FUNCTION "FC116_Inerting" : Void   // FC116, STL
{ S7_Optimized_Access := 'FALSE' }
AUTHOR : JaegerA
FAMILY : RS_KK
NAME : Inerting
VERSION : 1.1
   VAR_INPUT
      IN_Enable : Bool;
      IN_With_Inerting : Bool;   // Inerting selected in TP
      IN_OP_Mode_Manual : Bool;
      IN_OP_Mode_Wetshot : Bool;
      IN_OP_Mode_Test : Bool;
      IN_Start : Bool;
      IN_Stop : Bool;
      IN_T_Flushing : Bool;
      IN_T_Purge_Air : Bool;
      IN_Enable_pressurize_time : Bool;
      IN_AutoPurge_Air : Bool;
      IN_Quitt_Fault : Bool;
      IN_Cycle_runs : Bool;
      IN_MC_Activ : Bool;
      IN_PressurizeTimeRuns : Bool;
      IN_Shotend : Bool;
      IN_S_P_N2 : Bool;
      IN_S_P_FlushingAgent : Bool;
      IN_MH_selected : Bool;
      IN_Inert_MH : Bool;
      IN_Inert_Lance : Bool;
      IN_IntervalCleaning : Bool;
      IN_Ctrl_Fault_On : Bool;
      IN_Flowrate_N2_Actual : Real;
      IN_Shotwight : Real;
      IN_Foam_Density : DInt;
      IN_Leakage_value : Real;
      IN_DW_P_Build_Up_Before_Shot : S5Time;
      IN_DW_MaxInertTime : S5Time;
      IN_DW_Delay_Purge : S5Time;
      IN_DW_Ready_time : S5Time;
      IN_DW_Purge_time : S5Time;
      IN_DW_Delay_Plunger : S5Time;
      IN_DW_Delay_IntervalCleaning : S5Time;
      IN_DW_PurgeTime_IntervalCleaning : S5Time;
      IN_DW_PauseTime_IntervalCleaning : S5Time;
      IN_DW_Duration_IntervalCleaning : S5Time;
      IN_Timer_Delay_Leakage : Timer;
      IN_Timer_hourly_tact : Timer;
      IN_Timer_Inerting : Timer;
      IN_Timer_Ready : Timer;
      IN_Timer_Delay_Purge : Timer;
      IN_Timer_Purge : Timer;
      IN_Timer_Maximum_InertTime : Timer;
      IN_Timer_Delay_Plunger_N2 : Timer;
      IN_Timer_Delay_Tact : Timer;
      IN_Timer_PurgeTime_Tact : Timer;
      IN_Timer_PauseTime_Tact : Timer;
      IN_Timer_TotalTime_Tact : Timer;
   END_VAR
   VAR_OUTPUT
      OUT_H_Inert : Bool;
      OUT_H_Purge : Bool;
      OUT_H_FlushingAgent : Bool;
   END_VAR
   VAR_IN_OUT
      IO_DD_Inertfactor : Real;
      IO_DD_StartOffset : Real;
      IO_DD_DF_N2_SetValue : Real;
      IO_DD_DF_N2_Total : Real;
      IO_DD_DF_N2_Leakage : Real;
      IO_MH_Logged_on : Bool;
      IO_V_Piston : Bool;
      IO_V_Inert : Bool;
      IO_V_Purge_Air : Bool;
      IO_V_FlushingAgent : Bool;
      IO_Status : "UDT124_Inerting";   // Speichern der Antriebs- Zustände für das Programm
      IO_Status_Faults : "UDT1825_FLT_Inerting";
      IO_NewFault : Bool;
      IO_FaultLevel_1 : Bool;
      IO_FaultLevel_2 : Bool;
      IO_FaultLevel_3 : Bool;
   END_VAR
   VAR_TEMP
      Temp_IO_Status : "UDT124_Inerting";   // Temporärer Antriebs- Status für die interne Bearbeitung des Bausteins
      Temp_IO_Status_Faults : "UDT1825_FLT_Inerting";
      ERROR_CODE : Int;   // Störungszustand der Systemfunktion "BLKMOV" Blockmove
      Anyzeiger : ANY;   // Zeiger zum Kopieren der Bereiche "IO_Status" und "Temp_IO_Status"
      Anyzeiger2 : ANY;   // Zeiger zum Kopieren der Bereiche "IO_Status" und "Temp_IO_Status"
      InertTime : S5Time;
      Mem : Time;
      TimeValue : Word;
      Inertfactor : Int;
      Auto_Purge_On : Bool;
      Flag_StartTime : Bool;
      Hour_tact_ON : Bool;
      Quantity_N2_PressurizeTimeRuns : DInt;
      Total_Quantity_PressurizeTimeRuns : DInt;
      P_build_Up_time : DInt;
   END_VAR
BEGIN

REGION Network 1: Embed secured data
         LAR1;
         L;
         LAR2;
   //
         L     W#16#1002;  // Bytes
         T     W[AR1, P#0.0];
         L     6;  // Anzahl Bytes
         T     W[AR1, P#2.0];
         L     W[AR2, P#0.0];  // Baustein Nr.
         T     W[AR1, P#4.0];
         L     D[AR2, P#2.0];  // Datenanfang
         T     D[AR1, P#6.0];
   //
         CALL  BLKMOV
         ( SRCBLK  := #Anyzeiger,
           RET_VAL := #ERROR_CODE,
           DSTBLK  := #Temp_IO_Status
         );
   //
         LAR1;
         L;
         LAR2;
   //
         L     W#16#1002;  // Bytes
         T     W[AR1, P#0.0];
         L     2;  // Anzahl Bytes
         T     W[AR1, P#2.0];
         L     W[AR2, P#0.0];  // Baustein Nr.
         T     W[AR1, P#4.0];
         L     D[AR2, P#2.0];  // Datenanfang
         T     D[AR1, P#6.0];
   //
         CALL  BLKMOV
         ( SRCBLK  := #Anyzeiger2,
           RET_VAL := #ERROR_CODE,
           DSTBLK  := #Temp_IO_Status_Faults
         );
END_REGION

REGION Network 2: Faults
         CLR;
         =     #Temp_IO_Status.FaultLevel_1;
         =     #Temp_IO_Status.FaultLevel_2;
         =     #Temp_IO_Status.FaultLevel_3;
         =     #Temp_IO_Status.Message_activ;

   // Reset Faults
         A     #IN_Quitt_Fault;
         ON    #IN_With_Inerting;
         R     #Temp_IO_Status_Faults.Fault_P_N2;
         R     #Temp_IO_Status_Faults.Fault_flow_N2;
         R     #Temp_IO_Status_Faults.Fault_P_Flushing_Agent;
         R     #Temp_IO_Status_Faults.Fault_Leakage_N2;
         R     #Temp_IO_Status_Faults.Fault_MaxInertingTime;
         R     #Temp_IO_Status_Faults.Fault_NoShotwight;

   // Störung Vordruck N2
         AN    #IN_S_P_N2;
         A     #IN_Ctrl_Fault_On;
         A     #IN_MH_selected;
         A     #IN_With_Inerting;
         AN    #Temp_IO_Status_Faults.Fault_P_N2;
         S     #Temp_IO_Status_Faults.Fault_P_N2;
         S     #IO_NewFault;
   // Störung Vordruck Spülmittel
         A     #IN_MH_selected;
         A     #IN_With_Inerting;
         AN    #IN_S_P_FlushingAgent;
         AN    #Temp_IO_Status_Faults.Fault_P_Flushing_Agent;
         S     #Temp_IO_Status_Faults.Fault_P_Flushing_Agent;
         S     #IO_NewFault;
   // Störung Maximale Inertisierzeit überschritten
         A     #IO_V_Piston;
         A     #IN_With_Inerting;
         A     #Temp_IO_Status.Inert_runs;
         A     #IN_OP_Mode_Wetshot;
         A     #IN_Ctrl_Fault_On;
         A     #IN_MH_selected;
         L     #IN_DW_MaxInertTime;
         SD    #IN_Timer_Maximum_InertTime;
         A     #IN_Timer_Maximum_InertTime;
         AN    #Temp_IO_Status_Faults.Fault_MaxInertingTime;
         S     #Temp_IO_Status_Faults.Fault_MaxInertingTime;
         S     #IO_NewFault;

   // Störung Schussgewicht
         A     #IN_With_Inerting;
         A     #IN_Enable;
         A     #IN_Start;
         A     #IN_MH_selected;
         A(;
         L     #IN_Shotwight;
         L     0;
         ==D;
         );
         AN    #Temp_IO_Status_Faults.Fault_NoShotwight;
         S     #Temp_IO_Status_Faults.Fault_NoShotwight;
         S     #IO_NewFault;
END_REGION

REGION Network 3: Start and cancel
   // Start nur möglich wenn kein Zyklus läuft, denn es muß bei Zyklusstart die 
   // Schusszeit übertragen werden.
         A     #IN_Enable;
         A     #IN_Start;
         A     #IN_MH_selected;
         AN    #IN_Cycle_runs;
         AN    #Temp_IO_Status.OK;
         AN    #Temp_IO_Status_Faults.Fault_P_N2;
         AN    #Temp_IO_Status_Faults.Fault_flow_N2;
         AN    #Temp_IO_Status_Faults.Fault_NoShotwight;
         FP    #Temp_IO_Status.FH_Start;
         =     #Temp_IO_Status.FP_Start;

         A     #Temp_IO_Status.FP_Start;
         S     #Temp_IO_Status.Inert_started;

   // Abbruch
         ON    #IN_Enable;
         ON    #IN_Stop;
         ON    #IN_MH_selected;
         O     #Temp_IO_Status_Faults.Fault_P_N2;
         O     #Temp_IO_Status_Faults.Fault_flow_N2;
         O     #Temp_IO_Status_Faults.Fault_MaxInertingTime;
         O     #Temp_IO_Status.OK;
         R     #Temp_IO_Status.Inert_started;
         R     #Temp_IO_Status.Inert_runs;
         R     #Temp_IO_Status.FP_ST_received;
END_REGION

REGION Network 4: Calculate N2 flow
   // N² Spülmenge = Schussgewicht(g)/ Verschäumte Dichte PU (g/dm³) x Spülfaktor(1)
         L     #IO_DD_Inertfactor;
         L     8;
         >=D;
         JC    W1ok;
         L     8;
         T     #IO_DD_Inertfactor;

   W1ok: L     #IO_DD_StartOffset;
         L     0;
         >R;
         JC    W2ok;
         L     0;
         T     #IO_DD_StartOffset;

   W2ok: A     #Temp_IO_Status.Inert_started;
         FP    #Temp_IO_Status.FH_ST_received;
         S     #Temp_IO_Status.FP_ST_received;

         A     #Temp_IO_Status.FP_ST_received;
         JCN   ew;

         SET;
         S     #Temp_IO_Status.Inert_runs;

         L     #IN_Shotwight;
         L     #IN_Foam_Density;
         /D;
         L     #IO_DD_Inertfactor;
         *D;
         L     #IO_DD_StartOffset;
         +D;
         L     10;
         /D;
         T     #IO_DD_DF_N2_SetValue;

   ew:   NOP   0;
END_REGION

REGION Network 5: Inerting procedure start
         A     #Temp_IO_Status.Inert_runs;
         A     #IO_V_Piston;
         A     #Temp_IO_Status.Inert_runs;
         A(;
         L     #IO_DD_DF_N2_Total;
         L     #IO_DD_DF_N2_SetValue;
         >=D;
         );
         AN    #Temp_IO_Status_Faults.Fault_flow_N2;
         S     #Temp_IO_Status.OK;
         R     #Temp_IO_Status.Inert_runs;
END_REGION

REGION Network 6: Start PressurizeTimeRuns before Inerting is finished
         AN    #Temp_IO_Status.Inert_runs;
         O     #IN_Inert_Lance;
         ON    #IN_Enable_pressurize_time;
         R     #Temp_IO_Status.Start_PressurizeTimeRuns;
         JC    M001;

         CALL  "FC119_TConvert_ms"
         ( IN_S5_Time    := #IN_DW_P_Build_Up_Before_Shot,
           IN_Time_in_ms := #P_build_Up_time
         );

         L     #IN_Flowrate_N2_Actual;
         DTR;
         L     #P_build_Up_time;
         DTR;
         *R;
         L     1000.0;
         /R;
         RND;
         T     #Quantity_N2_PressurizeTimeRuns;

         L     #IO_DD_DF_N2_Total;
         L     #Quantity_N2_PressurizeTimeRuns;
         +D;
         T     #Total_Quantity_PressurizeTimeRuns;

         A(;
         L     #Total_Quantity_PressurizeTimeRuns;
         L     #IO_DD_DF_N2_SetValue;
         >=D;
         );
         A     #IO_V_Piston;
         =     #Temp_IO_Status.Start_PressurizeTimeRuns;
END_REGION

REGION Network 7: Start ready time, Start PressurizeTimeRuns
   M001: A     #Temp_IO_Status.OK;
         A     #IN_OP_Mode_Manual;
         L     #IN_DW_Ready_time;
         SD    #IN_Timer_Ready;

   // If Shot is not running, Reset ready time
         AN    #IN_Cycle_runs;
         O     #IN_PressurizeTimeRuns;
         A     #IN_Timer_Ready;
         O     #IN_Shotend;
         R     #Temp_IO_Status.Start_PressurizeTimeRuns;

         AN    #IN_Cycle_runs;
         A     #IN_Timer_Ready;
         O     #IN_Shotend;
         R     #Temp_IO_Status.OK;
END_REGION

REGION Network 8: Start Purge
         A     #IN_AutoPurge_Air;
         AN    #IN_OP_Mode_Test;
         A     #IN_Shotend;
         A     #IN_MH_selected;
         A(;
         L     #IN_DW_Purge_time;
         L     0;
         >I;
         );
         L     #IN_DW_Delay_Purge;
         SS    #IN_Timer_Delay_Purge;
         A     #IN_Timer_Delay_Purge;
         =     #Temp_IO_Status.Purge_runs;

         A     #Temp_IO_Status.Purge_runs;
         A     #IO_V_Piston;
         L     #IN_DW_Purge_time;
         SD    #IN_Timer_Purge;

         A     #IN_Timer_Purge;
         R     #Temp_IO_Status.Purge_runs;
         R     #IN_Timer_Purge;
         R     #IN_Timer_Delay_Purge;
END_REGION

REGION Network 9: Interval cleaning
         AN    #IN_IntervalCleaning;
         A     "DB619_State_MPart".Operationmode[1].Controllvoltage;
         JC    Vent;
         A     #Temp_IO_Status.Purge_runs;
         L     #IN_DW_Delay_IntervalCleaning;
         SF    #IN_Timer_Delay_Tact;

         A     #IN_Timer_Purge;
         O     #IN_Timer_Delay_Tact;
         FN    #Temp_IO_Status.FH_Start_Time;
         =     #Temp_IO_Status.FP_Start_Time;
         A     #Temp_IO_Status.FP_Start_Time;
         S     #Temp_IO_Status.FP_Start_Leakage_Control;

         A     #Temp_IO_Status.FP_Start_Time;
         L     #IN_DW_Duration_IntervalCleaning;
         SE    #IN_Timer_TotalTime_Tact;
         A     #IN_Timer_TotalTime_Tact;
         FN    #Temp_IO_Status.FH_Start_Leakage_Control;
         S     #Temp_IO_Status.Reserve26;

         AN    #IN_Timer_PauseTime_Tact;
         A     #IN_Timer_TotalTime_Tact;
         A     #IO_V_Piston;
         L     #IN_DW_PurgeTime_IntervalCleaning;
         SD    #IN_Timer_PurgeTime_Tact;
         A     #IN_Timer_PurgeTime_Tact;
         R     #Temp_IO_Status.FP_Start_Leakage_Control;

         A     #IN_Timer_PurgeTime_Tact;
         A     #IN_Timer_TotalTime_Tact;
         L     #IN_DW_PauseTime_IntervalCleaning;
         SE    #IN_Timer_PauseTime_Tact;
         A     #IN_Timer_PauseTime_Tact;
         FN    #Temp_IO_Status.FH_Start_Inert;
         A     #IN_Timer_TotalTime_Tact;
         S     #Temp_IO_Status.FP_Start_Leakage_Control;

         A     #IN_MC_Activ;
         O     #Temp_IO_Status.Inert_runs;
         O     #Temp_IO_Status.Reserve26;
         R     #IN_Timer_TotalTime_Tact;
         R     #IN_Timer_Delay_Tact;
         R     #Temp_IO_Status.FP_Start_Leakage_Control;
         R     #IN_Timer_PurgeTime_Tact;
         R     #IN_Timer_PauseTime_Tact;
         R     #Temp_IO_Status.Reserve26;

         JU    VENT_Mig;

   Vent: SET;
         R     #IN_Timer_TotalTime_Tact;
         R     #IN_Timer_Delay_Tact;
         R     #Temp_IO_Status.FP_Start_Leakage_Control;
         R     #Temp_IO_Status.Reserve26;
         R     #IN_Timer_PurgeTime_Tact;
         R     #IN_Timer_PauseTime_Tact;
END_REGION

REGION Network 10: Valves
   VENT_Mig:NOP   0;
   // Inertisieren bzw. Ausblasen
         A     #IO_V_Piston;  //#Temp_IO_Status.Inert_laeuft
         A     #IN_OP_Mode_Wetshot;
         AN    #Temp_IO_Status.Purge_runs;
         AN    #IN_T_Purge_Air;
         AN    #Temp_IO_Status.FP_Start_Leakage_Control;  // Taktausblasen
         =     #IO_V_Inert;

   // Spülen
         A     #IN_T_Flushing;
         AN    #IN_T_Purge_Air;
         AN    #IN_Cycle_runs;
         =     #IO_V_FlushingAgent;

   // Ausblasen Luft
         O     #Temp_IO_Status.Purge_runs;
         O     #IN_T_Purge_Air;
         O     #Temp_IO_Status.FP_Start_Leakage_Control;
         AN    #IN_T_Flushing;
   //    UN    #IN_Zyklus_laeuft
         =     #IO_V_Purge_Air;

   // Ventil Kolben
         O     #Temp_IO_Status.Inert_runs;
   //      O     #IO_V_Purge_Air      // Manuell beim Reinigen
         O     #IO_V_FlushingAgent;  // Manuell beim Spülen
         L     #IN_DW_Delay_Plunger;
         SD    #IN_Timer_Delay_Plunger_N2;
         A     #IN_Timer_Delay_Plunger_N2;
         O     #IO_V_Purge_Air;
         =     #IO_V_Piston;
END_REGION

REGION Network 11: Lamps
   // Inertisieren
         A(;
         AN    #IN_Cycle_runs;
         AN    #Temp_IO_Status.Inert_runs;
         A     #IN_OP_Mode_Wetshot;
         A     #IN_Enable;
         A     #IN_Stop;
         O;
         A     #Temp_IO_Status.Inert_runs;
         A     "Flag_01_250_Hertz";
         );

         A(;
         AN    #IN_Cycle_runs;
         AN    #Temp_IO_Status.OK;
         );
         =     #OUT_H_Inert;

   // Ausblasen N2 oder Luft
         A     #IO_V_Piston;
         AN    #IO_V_FlushingAgent;
         A     "Flag_01_250_Hertz";
         O     #IO_V_Purge_Air;
         =     #OUT_H_Purge;

   // Spülmittel
         A     #IO_V_FlushingAgent;
         =     #OUT_H_FlushingAgent;
END_REGION

REGION Network 12: If fault stop Inert
   // Inert bei STG abbrechen...
         O     #Temp_IO_Status_Faults.Fault_P_N2;
         O     #Temp_IO_Status_Faults.Fault_flow_N2;
         ON    #IN_Stop;
         R     #Temp_IO_Status.Inert_started;
         R     #Temp_IO_Status.Inert_runs;
         R     #Temp_IO_Status.Start_PressurizeTimeRuns;
         FP    #Temp_IO_Status.FH_Stop;
         =     #Temp_IO_Status.FP_Stop;
END_REGION

REGION Network 13: Leakage control
         AN    #Temp_IO_Status.Inert_started;
         L     S5T#15S;
         SD    #IN_Timer_Delay_Leakage;

         A     #Temp_IO_Status.Inert_started;
         O;
         A(;
         L     #IO_DD_DF_N2_Leakage;
         L     0;
         ==D;
         );
         R     #IN_Timer_hourly_tact;
         R     #Temp_IO_Status.Set_LoadValue;

         A     #Temp_IO_Status.Inert_started;
         JC    LE1;

         A     #IN_Timer_Delay_Leakage;
         AN    #IN_Timer_hourly_tact;
         =     #Hour_tact_ON;

   // Anstoss für das Laden des Zählers mit einem neuen Wert.
         A     #Hour_tact_ON;
         O;
         A     #Temp_IO_Status_Faults.Fault_Leakage_N2;
         FN    #Temp_IO_Status.Reserve27;
         S     #Temp_IO_Status.Set_LoadValue;

         A     #Hour_tact_ON;
         L     S5T#1H;
         SF    #IN_Timer_hourly_tact;

   // Wenn innerhalb des Stundentaktes der Leckageüberwachung der Zaehlwert erreicht wird,
   // dann wird eine Stoermeldung ausgegeben.
         A(;
         L     #IO_DD_DF_N2_Leakage;
         L     #IN_Leakage_value;
         >D;
         );
         AN    #Hour_tact_ON;
         A     #IN_Timer_hourly_tact;
         AN    #Temp_IO_Status.Set_LoadValue;
         S     #Temp_IO_Status_Faults.Fault_Leakage_N2;
         S     #IO_NewFault;

   LE1:  NOP   0;
END_REGION

REGION Network 14: Error handling
         O     #Temp_IO_Status_Faults.Fault_flow_N2;
         O     #Temp_IO_Status_Faults.Fault_MaxInertingTime;
         O     #Temp_IO_Status_Faults.Fault_NoShotwight;
         S     #Temp_IO_Status.FaultLevel_1;
         S     #IO_FaultLevel_1;

         O     #Temp_IO_Status_Faults.Fault_P_N2;
         S     #Temp_IO_Status.FaultLevel_2;
         S     #IO_FaultLevel_2;

         O     #Temp_IO_Status_Faults.Fault_P_Flushing_Agent;
         O     #Temp_IO_Status_Faults.Fault_MaxInertingTime;
         S     #Temp_IO_Status.FaultLevel_3;
         S     #IO_FaultLevel_3;
END_REGION

REGION Network 15: Save Datas
         CALL  BLKMOV
         ( SRCBLK  := #Temp_IO_Status,
           RET_VAL := #ERROR_CODE,
           DSTBLK  := #Anyzeiger
         );
   //
         CALL  BLKMOV
         ( SRCBLK  := #Temp_IO_Status_Faults,
           RET_VAL := #ERROR_CODE,
           DSTBLK  := #Anyzeiger2
         );
END_REGION
END_FUNCTION

FUNCTION "FC117_INT_Umwandler" : Void   // FC117, STL
{ S7_Optimized_Access := 'FALSE' }
VERSION : 0.1
BEGIN

REGION Network 1
   // Eingänge PU
         A     "DB119_Interface_Visu".APInterface[0].ExtP_OK;
         A     "DB119_Interface_Visu"."Inv.PrgNr";
         L     9;
         JC    m1;
         A     "DB119_Interface_Visu"."Inv.PrgNr";
         L     8;
         JC    m1;
         O     "DB119_Interface_Visu".Profibus;
         O     "DB119_Interface_Visu".Paritätsbit;
         A     "DB119_Interface_Visu".APInterface[0].ExtP_OK;
         L     7;
         JC    m1;
         O     "DB119_Interface_Visu".Paritätsbit;
         O     "DB119_Interface_Visu".Profibus;
         L     6;
   m1:   T     "Exp_Ok";

         A     "DB119_Interface_Visu".APInterface[0].Stop;
         A     "DB119_Interface_Visu"."Inv.PrgNr";
         L     7;
         JC    m6;
         A     "DB119_Interface_Visu"."Inv.PrgNr";
         L     6;
         JC    m6;
         O     "DB119_Interface_Visu".Profibus;
         O     "DB119_Interface_Visu".Paritätsbit;
         A     "DB119_Interface_Visu".APInterface[0].Stop;
         L     5;
         JC    m6;
         O     "DB119_Interface_Visu".Paritätsbit;
         O     "DB119_Interface_Visu".Profibus;
         L     4;
   m6:   T     "Stop";

         A     "DB119_Interface_Visu".APInterface[0].Strobe;
         A     "DB119_Interface_Visu"."Inv.PrgNr";
         L     5;
         JC    m2;
         A     "DB119_Interface_Visu"."Inv.PrgNr";
         L     4;
         JC    m2;
         O     "DB119_Interface_Visu".Profibus;
         O     "DB119_Interface_Visu".Paritätsbit;
         A     "DB119_Interface_Visu".APInterface[0].Strobe;
         L     3;
         JC    m2;
         O     "DB119_Interface_Visu".Paritätsbit;
         O     "DB119_Interface_Visu".Profibus;
         L     2;
   m2:   T     "Strobe";

         A     "DB119_Interface_Visu".APInterface[0].StrobeInv;
         AN    "DB119_Interface_Visu".Paritätsbit;
         L     3;
         JC    m3;
         A     "DB119_Interface_Visu".APInterface[0].StrobeInv;
         AN    "DB119_Interface_Visu".Paritätsbit;
         L     2;
         JC    m3;
         A     "DB119_Interface_Visu".APInterface[0].StrobeInv;
         A     "DB119_Interface_Visu".Paritätsbit;
         L     9;
         JC    m3;
         L     8;
   m3:   T     "StrobeInv";

         A     "DB119_Interface_Visu".APInterface[0].MH_open;
         L     1;
         JC    m4;
         L     0;
   m4:   T     "MH_open";
END_REGION

REGION Network 2
   // Ausgänge
         A     "DB119_Interface_Visu".APInterface[0].PU_OK;
         AN    "DB119_Interface_Visu".Profibus;
         L     11;
         JC    m7;
         AN    "DB119_Interface_Visu".Profibus;
         L     10;
         JC    m7;
         A     "DB119_Interface_Visu".APInterface[0].PU_OK;
         A     "DB119_Interface_Visu".Profibus;
         L     9;
         JC    m7;
         L     8;
   m7:   T     "PU_Ok";


         A     "DB119_Interface_Visu".APInterface[0].Strobe_quitt;
         L     9;
         JC    m10;
         L     8;
   m10:  T     "StrobeQuitt";

         A     "DB119_Interface_Visu".APInterface[0].cycle_run;
         L     7;
         JC    m11;
         L     6;
   m11:  T     "cycle_run";

         A     "DB119_Interface_Visu".APInterface[0].ready_for_shot;
         L     5;
         JC    m12;
         L     4;
   m12:  T     "ReadyForShot";

         A     "DB119_Interface_Visu".APInterface[0].shot_run;
         L     3;
         JC    m13;
         L     2;
   m13:  T     "ShotRun";

         A     "DB119_Interface_Visu".APInterface[0].shot_end;
         L     1;
         JC    m14;
         L     0;
   m14:  T     "ShotEnd";

         A     "DB119_Interface_Visu".APInterface[0].Service_mode;
         L     13;
         JC    m15;
         L     12;
   m15:  T     "ServiceMode";

         A     "DB119_Interface_Visu".APInterface[0].CP_is_forward;
         L     15;
         JC    m16;
         L     14;
   m16:  T     "CP_is_forward";
END_REGION
END_FUNCTION

FUNCTION "FC118_Enable_Inerting" : Void   // FC118, STL
{ S7_Optimized_Access := 'FALSE' }
VERSION : 0.1
   VAR_INPUT
      Prg_Number : Int;
      Ps_Number : Int;
      ReferenceValue : DInt;
   END_VAR
   VAR_OUTPUT
      Inerting_OFF : Bool;
      Shotwight : DInt;
   END_VAR
   VAR_TEMP
      PS_NR : Int;
      Startadress : Word;
      Offset : Word;
      Adress2 : Word;
      Toolnumber : Int;
   END_VAR
BEGIN

REGION Network 1
         L     #Prg_Number;  // Programmnummer
         L     2;
         *I;
         T     #Startadress;  // Anfangsadresse im Programm-DB
   ///
         L     #Startadress;  // Anfangsadresse im Programm-DB
         SLW   3;  // Adresse im DB
         T     #Startadress;  // Anfangsadresse im Programm-DB
         LAR2;  // in Adressregister 2 laden
   ///_____________________________________________________Werkzeug Nummer für Inertisierung
   //AUF   "DB940_Tool_alloc_automatic"
   //      L DBW [ AR2 , P#0.0 ]
   //      T     #Toolnumber
END_REGION

REGION Network 2
         A(;
         L     #Toolnumber;
         L     0;
         ==I;
         );
         O;
         A(;
         L     #Toolnumber;
         L     99;
         >I;
         );
         L     0;
         JC    M001;

         L     #Ps_Number;
         T     #PS_NR;

         L     #Toolnumber;  // Programmnummer
         L     416;
         *I;
         L     46;
         +I;
         T     #Startadress;  // Anfangsadresse im Programm-DB
         T     #Adress2;  // Für Schusszeiten
   ///
         L     #PS_NR;
         L     1;
         -I;
         L     52;
         *I;
         T     #Offset;

         L     #Startadress;  // Anfangsadresse im Programm-DB
         L     #Offset;
         +I;
         SLD   3;  // Adresse im DB
         T     #Startadress;  // Anfangsadresse im Programm-DB
         LAR2;  // in Adressregister 2 laden
   ///_____________________________________________________MK Nummer für Inertisierung
         OPN   "DB925_ShotData_1";
         L     DBD[AR2, P#0.0];
   M001: T     #Shotwight;
END_REGION

REGION Network 3
         L     #Shotwight;
         L     #ReferenceValue;
         <D;
         =     #Inerting_OFF;
END_REGION
END_FUNCTION

FUNCTION "FC119_TConvert_ms" : Void   // FC119, STL
TITLE = Konvertierung einer S5- Zeit in einen Milisekunden- Zeitwert
{ S7_Optimized_Access := 'FALSE' }
AUTHOR : KT242
FAMILY : RS_KK
NAME : TimConv
VERSION : 1.0
   VAR_INPUT
      IN_S5_Time : S5Time;   // Eingabe eines Zeitwertes im S5 Format
   END_VAR
   VAR_OUTPUT
      IN_Time_in_ms : DInt;   // Ausgabe des Zeitwertes in Millisekunden
   END_VAR
   VAR_TEMP
      Temp_Time_in_ms : DInt;
   END_VAR
BEGIN

REGION Network 1
         L     #IN_S5_Time;
         L     16#0FFF;
         AW;
         BTI;
         T     #IN_Time_in_ms;
         T     #Temp_Time_in_ms;
         L     #IN_S5_Time;
         L     16#3000;
         AW;
         SRW   12;
         JL    tban;  // case n
         JU    tba0;  // case 0
         JU    tba1;  // case 1
         JU    tba2;  // case 2
         JU    tba3;  // case 3
   tban: NOP   0;
   //
   tba0: L     10;  // 10ms
         L     #Temp_Time_in_ms;
         *D;
         T     #IN_Time_in_ms;
         JU    tbae;
   //
   tba1: L     100;  // 100ms
         L     #Temp_Time_in_ms;
         *D;
         T     #IN_Time_in_ms;
         JU    tbae;
   //
   tba2: L     1000;  // 1000ms
         L     #Temp_Time_in_ms;
         *D;
         T     #IN_Time_in_ms;
         JU    tbae;
   //
   tba3: L     10000;  // 10000ms
         L     #Temp_Time_in_ms;
         *D;
         T     #IN_Time_in_ms;
         JU    tbae;
   //
   tbae: NOP   0;
END_REGION
END_FUNCTION

FUNCTION "FC120_read_ProCan" : Void   // FC120, STL
TITLE = Read IO-Interface of ProCan modul
{ S7_Optimized_Access := 'FALSE' }
AUTHOR : KT242
FAMILY : RS_KK
NAME : RProcan
VERSION : 1.1
   VAR_TEMP
      Nullmerker : Byte;   // Zwischenmerker mit dem Wert "0" zum ablöschen bei gestörter Übertragung
      ERROR_CODE : Int;   // Störungszustand der Systemfunktion "FILL" Blockmove
      TempFlowState : Byte;
      Temp_InputSignals : DWord;
      dummy : Bool;
      TemRetBLKMOV : Int;
      TempMHStatus : Word;
      TempCPStatus : Byte;
      Temp_Einer : Word;
      Temp_Zehner : Word;
      Temp_QPBTime : S5Time;
   END_VAR
BEGIN

REGION Network 1: ProCan IO-Interface Flow 1
   //-------------------------------------------------------------------------------
   // Check, if PB-Module is accessible and without fault, otherwise do not
   // read data
   //-------------------------------------------------------------------------------
         AN    "PN_FlowRate".Component[1].FlowC_F.Active;
         JC    em01;

   //-----------------------------------------------------------------
   // Read address of flow component 01
   //-----------------------------------------------------------------
         L     "PN_FlowRate".Component[1].FlowC_F.Address;
         L     0;
         ==I;  //<>I
         JC    FLV1;
         L     "PN_FlowRate".Component[1].FlowC_F.Address;  // "DB1233_ProCanIO_Flow".AddressFlow[1].Ref_Act_FlowValue
   FLV1: T     "DB608_PV_Metering".Metering[1].Flow.PV_Conf_ActV.Address;

   //-----------------------------------------------------------------
   // Read state of flow component 1 and error handling component 1
   //-----------------------------------------------------------------
         L     "PN_FlowRate".Component[1].FlowC_F.Address;
         L     0;
         <=I;
         JC    FL01;
         L     "PN_FlowRate".Component[1].FlowC_F.Address;
         L     16;
         +D;
         SLD   3;
         LAR1;
         L     PIB [ AR1 , P#0.0 ];
   FL01: T     #TempFlowState;

   //------------------------------------------------------------------
   // Flow status
   //------------------------------------------------------------------
         CALL  BLKMOV
         ( SRCBLK  := #TempFlowState,
           RET_VAL := #TemRetBLKMOV,
           DSTBLK  := "DB122_FlowIndexState".MeteringUnit[1].IN_PROCAN.Flow_Status
         );

   //------------------------------------------------------------------
   // Flow status component 1 fault messages
   //------------------------------------------------------------------
         CALL  "FC054_FaultsMetering"
         ( IN_ProCanFlow_State := "DB122_FlowIndexState".MeteringUnit[1].IN_PROCAN.Flow_Status,  // #TempFlowState
           IN_Reset_Fault      := "DB009_Faults".Faults_Reset_FKT_M1,
           IO_Any_Flow_Fault   := "DB823_Error_Metering".MeteringPump[1],
           IO_HF_FLT_QPB       := "HF_FLT_QPB_C1",
           IO_FaultLevel1      := "DB009_Faults".Faults_FKT_Grp_1_M1,
           IO_FaultLevel2      := "DB009_Faults".Faults_FKT_Grp_2_M1,
           IO_FaultLevel3      := "DB009_Faults".Faults_FKT_Grp_3_M1,
           IO_NewFault         := "DB009_Faults".Faultschanging_M1
         );

         L     s5t#10s;
         T     #Temp_QPBTime;

         A     "DB122_FlowIndexState".MeteringUnit[1].IN_PROCAN.Flow_Status.FlowQPB;
         L     #Temp_QPBTime;
         SD    "TM_Alarm_QPBTime_C1";
         A     "TM_Alarm_QPBTime_C1";
         AN    "DB823_Error_Metering".MeteringPump[1].FLT_FlowSDATimeOut;
         S     "DB823_Error_Metering".MeteringPump[1].FLT_FlowSDATimeOut;
         S     "DB009_Faults".Faults_FKT_Grp_1_M1;
         S     "DB009_Faults".Faultschanging_M1;

   //------------------------------------------------------------------
   // Piston position
   //------------------------------------------------------------------
         L     "PN_FlowRate".Component[1].FlowC_F.Address;
         L     0;
         <>I;
         JC    PP01;
         L     "PN_FlowRate".Component[1].FlowC_F.Address;
         L     4;
         +D;
         SLD   3;
         LAR1;
         L     PID[AR1, P#0.0];
   PP01: T     "DB122_FlowIndexState".MeteringUnit[1].IN_PROCAN.PistonPosition;

   //------------------------------------------------------------------
   // Tandem status of piston 1, 2    (DB207 ???)
   //------------------------------------------------------------------
   //      L     "DB1233_ProCanIO_Flow".AddressFlow[1].Ref_TandemStatus
   //      L     0
   //      <=I
   //      SPB   PS01
   //      L     "DB1233_ProCanIO_Flow".AddressFlow[1].Ref_TandemStatus
   //      SLD   3
   //      LAR1
   //      L PEW [ AR1 , P#0.0 ]
   //PS01: T     "DB122_FlowIndexState".MeteringUnit[1].IN_PROCAN.TandemStatus
   //      T     %DB207.DBW0
   em01: NOP   0;
END_REGION

REGION Network 2: ProCan IO-Interface Flow 2
   //-------------------------------------------------------------------------------
   // Check, if PB-Module is accessible and without fault, otherwise do not
   // read data
   //-------------------------------------------------------------------------------
         AN    "PN_FlowRate".Component[2].FlowC_F.Active;
         JC    em02;

   //-----------------------------------------------------------------
   // Read address of flow component 01
   //-----------------------------------------------------------------
         L     "PN_FlowRate".Component[2].FlowC_F.Address;
         L     0;
         ==I;  //<>I
         JC    FLV2;
         L     "PN_FlowRate".Component[2].FlowC_F.Address;
   FLV2: T     "DB608_PV_Metering".Metering[2].Flow.PV_Conf_ActV.Address;

   //-----------------------------------------------------------------
   // Read state of flow component 1 and error handling component 1
   //-----------------------------------------------------------------
         L     "PN_FlowRate".Component[2].FlowC_F.Address;
         L     0;
         <=I;
         JC    FL02;
         L     "PN_FlowRate".Component[2].FlowC_F.Address;
         L     16;
         +D;
         SLD   3;
         LAR1;
         L     PIB [ AR1 , P#0.0 ];
   FL02: T     #TempFlowState;

   //-----------------------------------------------------------------
   // Transfer flowState
   //-----------------------------------------------------------------
         CALL  BLKMOV
         ( SRCBLK  := #TempFlowState,
           RET_VAL := #TemRetBLKMOV,
           DSTBLK  := "DB122_FlowIndexState".MeteringUnit[2].IN_PROCAN.Flow_Status
         );

   //------------------------------------------------------------------
   // Flow state component -> fault messages
   //------------------------------------------------------------------
         CALL  "FC054_FaultsMetering"
         ( IN_ProCanFlow_State := "DB122_FlowIndexState".MeteringUnit[2].IN_PROCAN.Flow_Status,
           IN_Reset_Fault      := "DB009_Faults".Faults_Reset_FKT_M1,
           IO_Any_Flow_Fault   := "DB823_Error_Metering".MeteringPump[2],
           IO_HF_FLT_QPB       := "HF_FLT_QPB_C2",
           IO_FaultLevel1      := "DB009_Faults".Faults_FKT_Grp_1_M1,
           IO_FaultLevel2      := "DB009_Faults".Faults_FKT_Grp_2_M1,
           IO_FaultLevel3      := "DB009_Faults".Faults_FKT_Grp_3_M1,
           IO_NewFault         := "DB009_Faults".Faultschanging_M1
         );

         A     "DB122_FlowIndexState".MeteringUnit[2].IN_PROCAN.Flow_Status.FlowQPB;
         L     #Temp_QPBTime;
         SD    "TM_Alarm_QPBTime_C2";
         A     "TM_Alarm_QPBTime_C2";
         AN    "DB823_Error_Metering".MeteringPump[2].FLT_FlowSDATimeOut;
         S     "DB823_Error_Metering".MeteringPump[2].FLT_FlowSDATimeOut;
         S     "DB009_Faults".Faults_FKT_Grp_1_M1;
         S     "DB009_Faults".Faultschanging_M1;

   //-----------------------------------------------------------------
   // Piston position
   //-----------------------------------------------------------------
         L     "PN_FlowRate".Component[2].FlowC_F.Address;
         L     0;
         <>I;
         JC    PP02;
         L     "PN_FlowRate".Component[2].FlowC_F.Address;
         L     4;
         +D;
         SLD   3;
         LAR1;
         L     PID[AR1, P#0.0];
   PP02: T     "DB122_FlowIndexState".MeteringUnit[2].IN_PROCAN.PistonPosition;

   //-----------------------------------------------------------------
   // Tandem state of Piston 3, 4
   //-----------------------------------------------------------------
   //      L     "DB1233_ProCanIO_Flow".AddressFlow[3].Ref_TandemStatus
   //      L     0
   //      <=I
   //      SPB   PS02
   //      L     "DB1233_ProCanIO_Flow".AddressFlow[3].Ref_TandemStatus
   //      SLD   3
   //      LAR1
   //      L PEW [ AR1 , P#0.0 ]
   //PS02: T     "DB122_FlowIndexState".MeteringUnit[2].IN_PROCAN.TandemStatus
   //      T     %DB207.DBW2
   em02: NOP   0;
END_REGION

REGION Network 3: ProCan IO-Interface flow 3
   //-------------------------------------------------------------------------------
   // Check, if PB-Modull is accessible and without fault, otherwithe do not
   // read data
   //-------------------------------------------------------------------------------
         AN    "PN_FlowRate".Component[3].FlowC_F.Active;
         JC    em03;

   //-----------------------------------------------------------------
   // Read address of flow component
   //-----------------------------------------------------------------
         L     "PN_FlowRate".Component[3].FlowC_F.Address;
         L     0;
         ==I;  //<>I
         JC    FLV3;
         L     "PN_FlowRate".Component[3].FlowC_F.Address;
   FLV3: T     "DB608_PV_Metering".Metering[3].Flow.PV_Conf_ActV.Address;

   //-----------------------------------------------------------------
   // Read state of flow component and error handling component
   //-----------------------------------------------------------------
         L     "PN_FlowRate".Component[3].FlowC_F.Address;
         L     0;
         <=I;
         JC    FL03;
         L     "PN_FlowRate".Component[3].FlowC_F.Address;
         L     16;
         +D;
         SLD   3;
         LAR1;
         L     PIB [ AR1 , P#0.0 ];
   FL03: T     #TempFlowState;

   //-----------------------------------------------------------------
   // Transfer flowState
   //-----------------------------------------------------------------
         CALL  BLKMOV
         ( SRCBLK  := #TempFlowState,
           RET_VAL := #TemRetBLKMOV,
           DSTBLK  := "DB122_FlowIndexState".MeteringUnit[3].IN_PROCAN.Flow_Status
         );

   //------------------------------------------------------------------
   // Flow state component -> fault messages
   //------------------------------------------------------------------
         CALL  "FC054_FaultsMetering"
         ( IN_ProCanFlow_State := "DB122_FlowIndexState".MeteringUnit[3].IN_PROCAN.Flow_Status,
           IN_Reset_Fault      := "DB009_Faults".Faults_Reset_FKT_M1,
           IO_Any_Flow_Fault   := "DB823_Error_Metering".MeteringPump[3],
           IO_HF_FLT_QPB       := "HF_FLT_QPB_C3",
           IO_FaultLevel1      := "DB009_Faults".Faults_FKT_Grp_1_M1,
           IO_FaultLevel2      := "DB009_Faults".Faults_FKT_Grp_2_M1,
           IO_FaultLevel3      := "DB009_Faults".Faults_FKT_Grp_3_M1,
           IO_NewFault         := "DB009_Faults".Faultschanging_M1
         );

   //-----------------------------------------------------------------
   // Piston position
   //-----------------------------------------------------------------
         L     "PN_FlowRate".Component[3].FlowC_F.Address;
         L     0;
         <>I;
         JC    PP03;
         L     "PN_FlowRate".Component[3].FlowC_F.Address;
         L     4;
         +D;
         SLD   3;
         LAR1;
         L     PID[AR1, P#0.0];
   PP03: T     "DB122_FlowIndexState".MeteringUnit[3].IN_PROCAN.PistonPosition;

   //-----------------------------------------------------------------
   // Tandem state of Piston 5, 6
   //-----------------------------------------------------------------
   //      L     "DB1233_ProCanIO_Flow".AddressFlow[5].Ref_TandemStatus
   //      L     0
   //      <=I
   //      SPB   PS03
   //      L     "DB1233_ProCanIO_Flow".AddressFlow[5].Ref_TandemStatus
   //      SLD   3
   //      LAR1
   //      L PEW [ AR1 , P#0.0 ]
   //PS03: T     "DB122_FlowIndexState".MeteringUnit[3].IN_PROCAN.TandemStatus
   //      T     %DB207.DBW2
   em03: NOP   0;
END_REGION

REGION Network 4: ProCan IO-Interface flow 4
   //-------------------------------------------------------------------------------
   // Check, if PB-Modull is accessible and without fault, otherwithe do not
   // read data
   //-------------------------------------------------------------------------------
         AN    "PN_FlowRate".Component[4].FlowC_F.Active;
         JC    em04;

   //-----------------------------------------------------------------
   // Read address of flow component
   //-----------------------------------------------------------------
         L     "PN_FlowRate".Component[4].FlowC_F.Address;
         L     0;
         ==I;  //<>I
         JC    FLV4;
         L     "PN_FlowRate".Component[4].FlowC_F.Address;
   FLV4: T     "DB608_PV_Metering".Metering[4].Flow.PV_Conf_ActV.Address;

   //-----------------------------------------------------------------
   // Read state of flow component and error handling component
   //-----------------------------------------------------------------
         L     "PN_FlowRate".Component[4].FlowC_F.Address;
         L     0;
         <=I;
         JC    FL04;
         L     "PN_FlowRate".Component[4].FlowC_F.Address;
         L     16;
         +D;
         SLD   3;
         LAR1;
         L     PIB [ AR1 , P#0.0 ];
   FL04: T     #TempFlowState;

   //-----------------------------------------------------------------
   // Transfer flowState
   //-----------------------------------------------------------------
         CALL  BLKMOV
         ( SRCBLK  := #TempFlowState,
           RET_VAL := #TemRetBLKMOV,
           DSTBLK  := "DB122_FlowIndexState".MeteringUnit[4].IN_PROCAN.Flow_Status
         );

   //------------------------------------------------------------------
   // Flow state component -> fault messages
   //------------------------------------------------------------------
         CALL  "FC054_FaultsMetering"
         ( IN_ProCanFlow_State := "DB122_FlowIndexState".MeteringUnit[4].IN_PROCAN.Flow_Status,
           IN_Reset_Fault      := "DB009_Faults".Faults_Reset_FKT_M1,
           IO_Any_Flow_Fault   := "DB823_Error_Metering".MeteringPump[4],
           IO_HF_FLT_QPB       := "HF_FLT_QPB_C4",
           IO_FaultLevel1      := "DB009_Faults".Faults_FKT_Grp_1_M1,
           IO_FaultLevel2      := "DB009_Faults".Faults_FKT_Grp_2_M1,
           IO_FaultLevel3      := "DB009_Faults".Faults_FKT_Grp_3_M1,
           IO_NewFault         := "DB009_Faults".Faultschanging_M1
         );

   //-----------------------------------------------------------------
   // Piston position
   //-----------------------------------------------------------------
         L     "PN_FlowRate".Component[4].FlowC_F.Address;
         L     0;
         <>I;
         JC    PP04;
         L     "PN_FlowRate".Component[4].FlowC_F.Address;
         L     4;
         +D;
         SLD   3;
         LAR1;
         L     PID[AR1, P#0.0];
   PP04: T     "DB122_FlowIndexState".MeteringUnit[4].IN_PROCAN.PistonPosition;

   //-----------------------------------------------------------------
   // Tandem state of Piston 7,8
   //-----------------------------------------------------------------
   //      L     "DB1233_ProCanIO_Flow".AddressFlow[7].Ref_TandemStatus
   //      L     0
   //      <=I
   //      SPB   PS04
   //      L     "DB1233_ProCanIO_Flow".AddressFlow[7].Ref_TandemStatus
   //      SLD   3
   //      LAR1
   //      L PEW [ AR1 , P#0.0 ]
   //PS04: T     "DB122_FlowIndexState".MeteringUnit[4].IN_PROCAN.TandemStatus
   //      T     %DB207.DBW2
   em04: NOP   0;
END_REGION

REGION Network 5: Mixing head IO-Interface of mixing head 1
   //----------------------------------------------------------------
   // Check if ProfiBus member is accessible and without fault
   // otherwise no communication is possible
   //----------------------------------------------------------------
         A     "PN_Mixinghead".Mixinghead[1].Digital.Active;
         JC    mk1;
         L     0;
         T     #Nullmerker;
         CALL  FILL
         ( BVAL    := #Nullmerker,
           RET_VAL := #ERROR_CODE,
           BLK     := "DB123_MH_IO_Signals".MH[1]
         );
         JU    emk1;
   //_________________________________________________________________
   //
   mk1:  NOP   0;
   // Digital Input -> Ini Signals mixinghead, cleaningpiston

         A     "ES_OP_Panel_MH01";
         =     "DB123_MH_IO_Signals".MH[1].IN.MH_EmergencyStop;
         A     "IPS_CP_MH01";
         =     "DB123_MH_IO_Signals".MH[1].IN.MH_APS_CleaningPiston;
         A     "S_Rel_SWU_MH01";
         =     "DB123_MH_IO_Signals".MH[1].IN.MH_Release_SWU;
         A     "S_Manuel_MH01";
         =     "DB123_MH_IO_Signals".MH[1].IN.MH_Manual_Mode;
         A     "S_Automatic_MH01";
         =     "DB123_MH_IO_Signals".MH[1].IN.MH_Auto_Mode;

         O     "K_PreparationFoamingMC01";
         =     "DB123_MH_IO_Signals".MH[1].IN.MH_Prep_Foaming_MC;
         O     "K_FoamingReleaseMC01";
         =     "DB123_MH_IO_Signals".MH[1].IN.MH_Releas_Foaming_MC;
   ///
         L     "S_ProgNoSelectMH01";
         AW    16#000F;
         T     "DB123_MH_IO_Signals".MH[1].IN.MH_Prog_No_MH;

         AN    "DB704_MH_Value".Mixinghead[1].With99program;
         JC    No99Prog;
         L     "S_ProgNoSelectMH01";
         L     16#0f;
         AW;
         T     #Temp_Einer;  // Zwischenspeichern Einer
   //
         L     0;
         T     #Temp_Zehner;
   //-
         AN    "S_ProgrNo_Bit10_MH01";
         JC    noValue10;
         +     10;
   noValue10:NOP   0;

         AN    "S_ProgrNo_Bit20_MH01";
         JC    noValue20;
         +     20;
   noValue20:NOP   0;

         AN    "S_ProgrNo_Bit40_MH01";
         JC    noValue40;
         +     40;
   noValue40:NOP   0;

         AN    "S_ProgrNo_Bit80_MH01";
         JC    noValue80;
         +     80;
   noValue80:NOP   0;

         L     #Temp_Einer;
         +I;
         T     "DB123_MH_IO_Signals".MH[1].IN.MH_Prog_No_MH;
   No99Prog:NOP   0;
         A     "T_Highpressure_MH01";
         =     "DB123_MH_IO_Signals".MH[1].IN.MH_HP_Circ_MH;
         A     "T_Start_MH01";
         =     "DB123_MH_IO_Signals".MH[1].IN.MH_Start;
         A     "T_Stop_MH01";
         =     "DB123_MH_IO_Signals".MH[1].IN.MH_Stop;
         A     "T_CP_forward_MH01";
         =     "DB123_MH_IO_Signals".MH[1].IN.MH_CP_forward;
         A     "T_CP_back_MH01";
         =     "DB123_MH_IO_Signals".MH[1].IN.MH_CP_backward;
         A     "IPS_MH_MH01";
         =     "DB123_MH_IO_Signals".MH[1].IN.MH_Aps_Mixinghead;

   MHS1: NOP   0;
   //-----------------------------------------------------------------
   // Shot status of MH-01
   //-----------------------------------------------------------------
         L     "PN_Mixinghead".Mixinghead[1].Digital.Address;
         L     0;
         ==D;
         JC    MS01;
         L     "PN_Mixinghead".Mixinghead[1].Digital.Address;
         L     12;
         +D;
         SLD   3;
         LAR1;
         L     PIW [ AR1 , P#0.0 ];
   MS01: T     #TempMHStatus;  // ProCan-MH_Status MH01

         CALL  BLKMOV
         ( SRCBLK  := #TempMHStatus,
           RET_VAL := #TemRetBLKMOV,
           DSTBLK  := "DB123_MH_IO_Signals".MH[1].IN.MH_Status
         );

   //
   //-----------------------------------------------------------------
   // Status of cleaning piston MH-01
   //-----------------------------------------------------------------
         A(;
         L     "PN_Mixinghead".Mixinghead[1].ReinigungskolbenDigital.Address;
         L     0;
         ==D;
         );
         ON    "PN_Mixinghead".Mixinghead[1].ReinigungskolbenDigital.Active;
         JC    CP01;
         L     "PN_Mixinghead".Mixinghead[1].ReinigungskolbenDigital.Address;
         L     8;
         +D;
         SLD   3;
         LAR1;
         L     PIB [ AR1 , P#0.0 ];
   CP01: T     #TempCPStatus;

         CALL  BLKMOV
         ( SRCBLK  := #TempCPStatus,
           RET_VAL := #TemRetBLKMOV,
           DSTBLK  := "DB123_MH_IO_Signals".MH[1].IN.CleaningPistonState
         );

   //-----------------------------------------------------------------
   // Actual shot time of MH-01
   //-----------------------------------------------------------------
         L     "PN_Mixinghead".Mixinghead[1].Digital.Address;
         L     0;
         ==D;
         JC    ST01;

         L     "PN_Mixinghead".Mixinghead[1].Digital.Address;
         SLD   3;
         LAR1;
         L     PID[AR1, P#0.0];
   ST01: T     "DB123_MH_IO_Signals".MH[1].IN.Shottime;

         AN    "DB123_MH_IO_Signals".MH[1].IN.MH_Status.shotdone_MH;
         JC    ShD1;

         L     "PN_Mixinghead".Mixinghead[1].Digital.Address;
         L     4;
         +D;
         SLD   3;
         LAR1;
         L     PID [ AR1 , P#0.0 ];
         T     "DB123_MH_IO_Signals".MH[1].IN.MH_Opentime;

         L     "PN_Mixinghead".Mixinghead[1].Digital.Address;
         L     8;
         +D;
         SLD   3;
         LAR1;
         L     PID [ AR1 , P#0.0 ];
         T     "DB123_MH_IO_Signals".MH[1].IN.MH_Closingtime;
   ShD1: NOP   0;
   emk1: NOP   0;
END_REGION

REGION Network 6: Read ProCan Data of MH-02
   //----------------------------------------------------------------
   // Check if ProfiBus member is accessible and without fault
   // otherwise no communication is possible
   //----------------------------------------------------------------
         A     "PN_Mixinghead".Mixinghead[2].Digital.Active;
         JC    mk2;
         L     0;
         T     #Nullmerker;
         CALL  FILL
         ( BVAL    := #Nullmerker,
           RET_VAL := #ERROR_CODE,
           BLK     := "DB123_MH_IO_Signals".MH[2]
         );
         JU    emk2;
   //_________________________________________________________________
   //
   mk2:  NOP   0;
   // Digital Input -> Ini Signals mixinghead, cleaningpiston

         A     "ES_OP_Panel_MH02";
         =     "DB123_MH_IO_Signals".MH[2].IN.MH_EmergencyStop;
         A     "IPS_CP_MH02";
         =     "DB123_MH_IO_Signals".MH[2].IN.MH_APS_CleaningPiston;
         SET;
         =     "DB123_MH_IO_Signals".MH[2].IN.MH_With_CleaningPiston;
         A     "S_Rel_SWU_MH02";
         =     "DB123_MH_IO_Signals".MH[2].IN.MH_Release_SWU;
         A     "S_Manuel_MH02";
         =     "DB123_MH_IO_Signals".MH[2].IN.MH_Manual_Mode;
         A     "S_Automatic_MH02";
         =     "DB123_MH_IO_Signals".MH[2].IN.MH_Auto_Mode;

         O     "K_PreparationFoamingMC02";
         =     "DB123_MH_IO_Signals".MH[2].IN.MH_Prep_Foaming_MC;
         O     "K_FoamingReleaseMC02";
         =     "DB123_MH_IO_Signals".MH[2].IN.MH_Releas_Foaming_MC;
   ///
         L     "S_ProgNoSelectMH02";
         AW    16#000F;
         T     #Temp_Einer;
   //
   //      L     "S_ProgNoSelectMH02"
   //      UW    16#000F
   //      L     10
   //      *I
   //      L     #Temp_Einer
   //      +I
         T     "DB123_MH_IO_Signals".MH[2].IN.MH_Prog_No_MH;